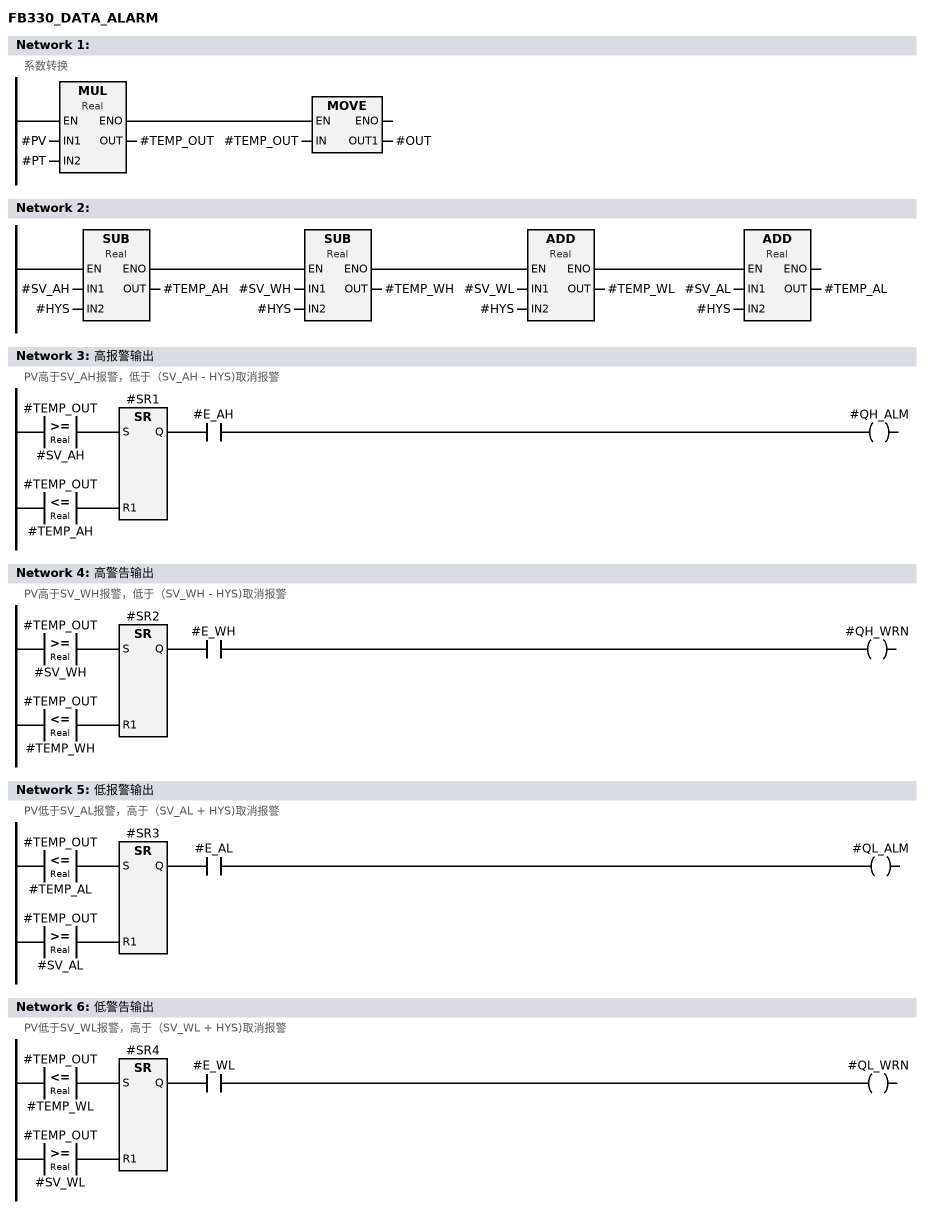
   RUNG wire#powerrail
      { S7_Templates := "SrcType := Real"; S7_GenerateENO := "TRUE" } Mul(in1 := #PV, in2 := #PT, out => #TEMP_OUT)
      { S7_GenerateENO := "TRUE" } Move(in := #TEMP_OUT, out1 => #OUT)
   END_RUNG
   // the same network as SCL:
   // ENO of a box is taken as its EN; it also drops when the box reports an error
   #TEMP_OUT := #PV * #PT;
   #OUT := #TEMP_OUT;
END_REGION

REGION Network 2
   RUNG wire#powerrail
      { S7_Templates := "SrcType := Real"; S7_GenerateENO := "TRUE" } Sub(in1 := #SV_AH, in2 := #HYS, out => #TEMP_AH)
      { S7_Templates := "SrcType := Real"; S7_GenerateENO := "TRUE" } Sub(in1 := #SV_WH, in2 := #HYS, out => #TEMP_WH)
      { S7_Templates := "SrcType := Real"; S7_GenerateENO := "TRUE" } Add(in1 := #SV_WL, in2 := #HYS, out => #TEMP_WL)
      { S7_Templates := "SrcType := Real"; S7_GenerateENO := "TRUE" } Add(in1 := #SV_AL, in2 := #HYS, out => #TEMP_AL)
   END_RUNG
   // the same network as SCL:
   // ENO of a box is taken as its EN; it also drops when the box reports an error
   #TEMP_AH := #SV_AH - #HYS;
   #TEMP_WH := #SV_WH - #HYS;
   #TEMP_WL := #SV_WL + #HYS;
   #TEMP_AL := #SV_AL + #HYS;
END_REGION

REGION Network 3: 高报警输出
   // PV高于SV_AH报警，低于（SV_AH - HYS)取消报警
   RUNG wire#powerrail
      { S7_Templates := "SrcType := Real" } GE_Contact(in1 := #TEMP_OUT, in2 := #SV_AH)
      S_SR(operand := #SR1, r1 := wire#w1)
      Contact( #E_AH )
      Coil( #QH_ALM )
   END_RUNG
   RUNG wire#powerrail
      { S7_Templates := "SrcType := Real" } LE_Contact(in1 := #TEMP_OUT, in2 := #TEMP_AH)
   END_RUNG wire#w1
   // the same network as SCL:
   IF #TEMP_OUT >= #SV_AH THEN
       #SR1 := TRUE;   // SR flip-flop
   END_IF;
   IF #TEMP_OUT <= #TEMP_AH THEN #SR1 := FALSE; END_IF;
   #QH_ALM := #SR1 AND #E_AH;
END_REGION

REGION Network 4: 高警告输出
   // PV高于SV_WH报警，低于（SV_WH - HYS)取消报警
   RUNG wire#powerrail
      { S7_Templates := "SrcType := Real" } GE_Contact(in1 := #TEMP_OUT, in2 := #SV_WH)
      S_SR(operand := #SR2, r1 := wire#w1)
      Contact( #E_WH )
      Coil( #QH_WRN )
   END_RUNG
   RUNG wire#powerrail
      { S7_Templates := "SrcType := Real" } LE_Contact(in1 := #TEMP_OUT, in2 := #TEMP_WH)
   END_RUNG wire#w1
   // the same network as SCL:
   IF #TEMP_OUT >= #SV_WH THEN
       #SR2 := TRUE;   // SR flip-flop
   END_IF;
   IF #TEMP_OUT <= #TEMP_WH THEN #SR2 := FALSE; END_IF;
   #QH_WRN := #SR2 AND #E_WH;
END_REGION

REGION Network 5: 低报警输出
   // PV低于SV_AL报警，高于（SV_AL + HYS)取消报警
   RUNG wire#powerrail
      { S7_Templates := "SrcType := Real" } LE_Contact(in1 := #TEMP_OUT, in2 := #TEMP_AL)
      S_SR(operand := #SR3, r1 := wire#w1)
      Contact( #E_AL )
      Coil( #QL_ALM )
   END_RUNG
   RUNG wire#powerrail
      { S7_Templates := "SrcType := Real" } GE_Contact(in1 := #TEMP_OUT, in2 := #SV_AL)
   END_RUNG wire#w1
   // the same network as SCL:
   IF #TEMP_OUT <= #TEMP_AL THEN
       #SR3 := TRUE;   // SR flip-flop
   END_IF;
   IF #TEMP_OUT >= #SV_AL THEN #SR3 := FALSE; END_IF;
   #QL_ALM := #SR3 AND #E_AL;
END_REGION

REGION Network 6: 低警告输出
   // PV低于SV_WL报警，高于（SV_WL + HYS)取消报警
   RUNG wire#powerrail
      { S7_Templates := "SrcType := Real" } LE_Contact(in1 := #TEMP_OUT, in2 := #TEMP_WL)
      S_SR(operand := #SR4, r1 := wire#w1)
      Contact( #E_WL )
      Coil( #QL_WRN )
   END_RUNG
   RUNG wire#powerrail
      { S7_Templates := "SrcType := Real" } GE_Contact(in1 := #TEMP_OUT, in2 := #SV_WL)
   END_RUNG wire#w1
   // the same network as SCL:
   IF #TEMP_OUT <= #TEMP_WL THEN
       #SR4 := TRUE;   // SR flip-flop
   END_IF;
   IF #TEMP_OUT >= #SV_WL THEN #SR4 := FALSE; END_IF;
   #QL_WRN := #SR4 AND #E_WL;
END_REGION
END_FUNCTION_BLOCK

FUNCTION "电机控制" : Void   // FC1, LAD
{ S7_Optimized_Access := 'FALSE' }
VERSION : 0.1
   VAR_TEMP   // added for the SCL form of the ladder/FBD networks
      _w1 : Bool;
      _s5time1 : S5Time;
      _w2 : Bool;
   END_VAR
BEGIN

REGION Network 1
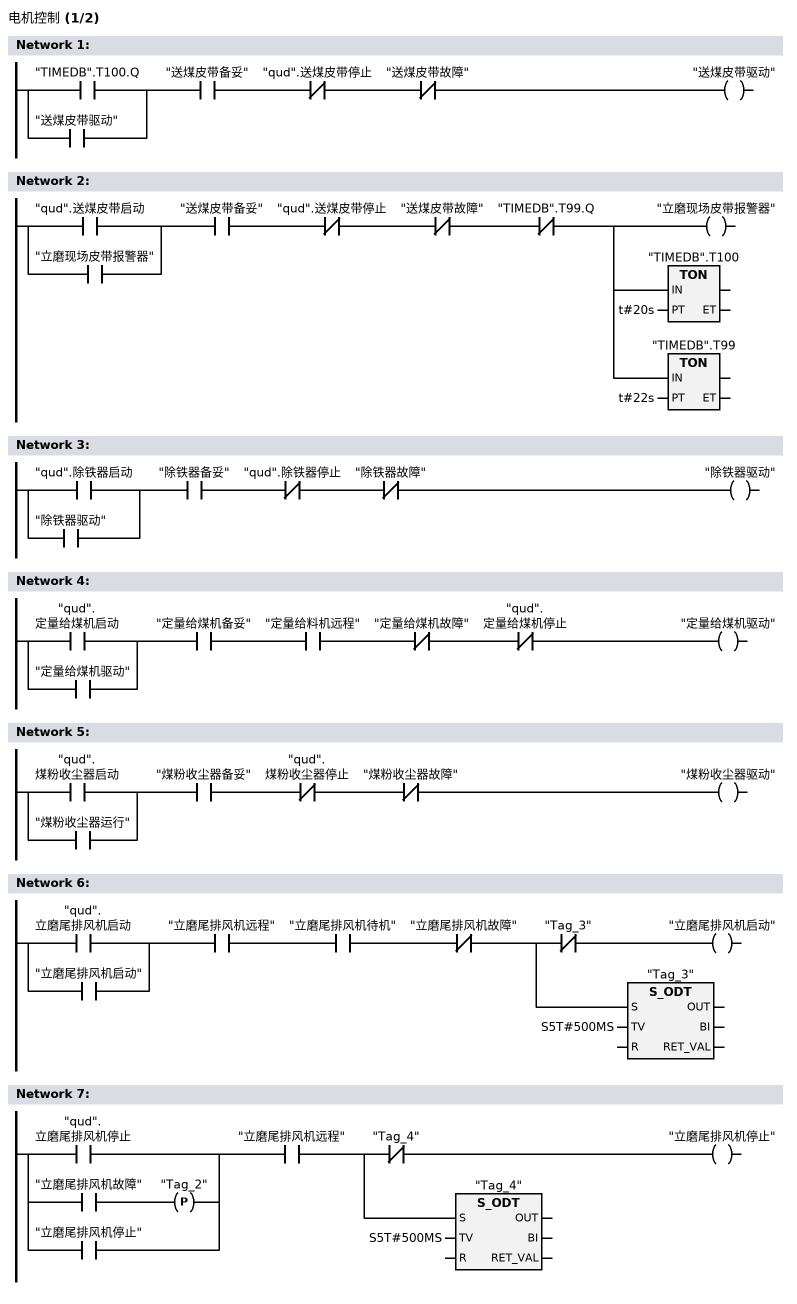
   RUNG wire#powerrail
      Contact( "TIMEDB".T100.Q )
      wire#w1
      Contact( "送煤皮带备妥" )
      I_Contact( "qud".送煤皮带停止 )
      I_Contact( "送煤皮带故障" )
      Coil( "送煤皮带驱动" )
   END_RUNG
   RUNG wire#powerrail
      Contact( "送煤皮带驱动" )
   END_RUNG wire#w1
   // the same network as SCL:
   "送煤皮带驱动" := ("TIMEDB".T100.Q OR "送煤皮带驱动") AND "送煤皮带备妥" AND NOT "qud".送煤皮带停止 AND NOT "送煤皮带故障";
END_REGION

REGION Network 2
   "立磨现场皮带报警器" := ("qud".送煤皮带启动 OR "立磨现场皮带报警器") AND "送煤皮带备妥" AND NOT "qud".送煤皮带停止 AND NOT "送煤皮带故障" AND NOT "TIMEDB".T99.Q;
   "TIMEDB".T100.TON(IN := "立磨现场皮带报警器", PT := t#20s);
   "TIMEDB".T99.TON(IN := "立磨现场皮带报警器", PT := t#22s);
END_REGION

REGION Network 3
   RUNG wire#powerrail
      Contact( "qud".除铁器启动 )
      wire#w1
      Contact( "除铁器备妥" )
      I_Contact( "qud".除铁器停止 )
      I_Contact( "除铁器故障" )
      Coil( "除铁器驱动" )
   END_RUNG
   RUNG wire#powerrail
      Contact( "除铁器驱动" )
   END_RUNG wire#w1
   // the same network as SCL:
   "除铁器驱动" := ("qud".除铁器启动 OR "除铁器驱动") AND "除铁器备妥" AND NOT "qud".除铁器停止 AND NOT "除铁器故障";
END_REGION

REGION Network 4
   RUNG wire#powerrail
      Contact( "qud".定量给煤机启动 )
      wire#w1
      Contact( "定量给煤机备妥" )
      Contact( "定量给料机远程" )
      I_Contact( "定量给煤机故障" )
      I_Contact( "qud".定量给煤机停止 )
      Coil( "定量给煤机驱动" )
   END_RUNG
   RUNG wire#powerrail
      Contact( "定量给煤机驱动" )
   END_RUNG wire#w1
   // the same network as SCL:
   "定量给煤机驱动" := ("qud".定量给煤机启动 OR "定量给煤机驱动") AND "定量给煤机备妥" AND "定量给料机远程" AND NOT "定量给煤机故障" AND NOT "qud".定量给煤机停止;
END_REGION

REGION Network 5
   RUNG wire#powerrail
      Contact( "qud".煤粉收尘器启动 )
      wire#w1
      Contact( "煤粉收尘器备妥" )
      I_Contact( "qud".煤粉收尘器停止 )
      I_Contact( "煤粉收尘器故障" )
      Coil( "煤粉收尘器驱动" )
   END_RUNG
   RUNG wire#powerrail
      Contact( "煤粉收尘器运行" )
   END_RUNG wire#w1
   // the same network as SCL:
   "煤粉收尘器驱动" := ("qud".煤粉收尘器启动 OR "煤粉收尘器运行") AND "煤粉收尘器备妥" AND NOT "qud".煤粉收尘器停止 AND NOT "煤粉收尘器故障";
END_REGION

REGION Network 6
   RUNG wire#powerrail
      Contact( "qud".立磨尾排风机启动 )
      wire#w1
      Contact( "立磨尾排风机远程" )
      Contact( "立磨尾排风机待机" )
      I_Contact( "立磨尾排风机故障" )
      wire#w2
      I_Contact( "Tag_3" )
      Coil( "立磨尾排风机启动" )
   END_RUNG
   RUNG wire#powerrail
      Contact( "立磨尾排风机启动" )
   END_RUNG wire#w1
   RUNG wire#w2
      S_ODT(T_NO := "Tag_3", TV := S5T#500MS, R :=, BI =>, RET_VAL =>)
   END_RUNG
   // the same network as SCL:
   #_w1 := ("qud".立磨尾排风机启动 OR "立磨尾排风机启动") AND "立磨尾排风机远程" AND "立磨尾排风机待机" AND NOT "立磨尾排风机故障";
   "立磨尾排风机启动" := #_w1 AND NOT "Tag_3";
   #_s5time1 := S_ODT(T_NO := "Tag_3", S := #_w1, TV := S5T#500MS);
END_REGION

REGION Network 7
   RUNG wire#powerrail
      Contact( "qud".立磨尾排风机停止 )
      wire#w1
      Contact( "立磨尾排风机远程" )
      wire#w2
      I_Contact( "Tag_4" )
      Coil( "立磨尾排风机停止" )
   END_RUNG
   RUNG wire#powerrail
      Contact( "立磨尾排风机故障" )
      P_Trig( "Tag_2" )
   END_RUNG wire#w1
   RUNG wire#powerrail
      Contact( "立磨尾排风机停止" )
   END_RUNG wire#w1
   RUNG wire#w2
      S_ODT(T_NO := "Tag_4", TV := S5T#500MS, R :=, BI =>, RET_VAL =>)
   END_RUNG
   // the same network as SCL:
   #_w1 := "立磨尾排风机故障" AND NOT "Tag_2";   // rising edge
   "Tag_2" := "立磨尾排风机故障";
   #_w2 := ("qud".立磨尾排风机停止 OR #_w1 OR "立磨尾排风机停止") AND "立磨尾排风机远程";
   "立磨尾排风机停止" := #_w2 AND NOT "Tag_4";
   #_s5time1 := S_ODT(T_NO := "Tag_4", S := #_w2, TV := S5T#500MS);
END_REGION

REGION Network 8
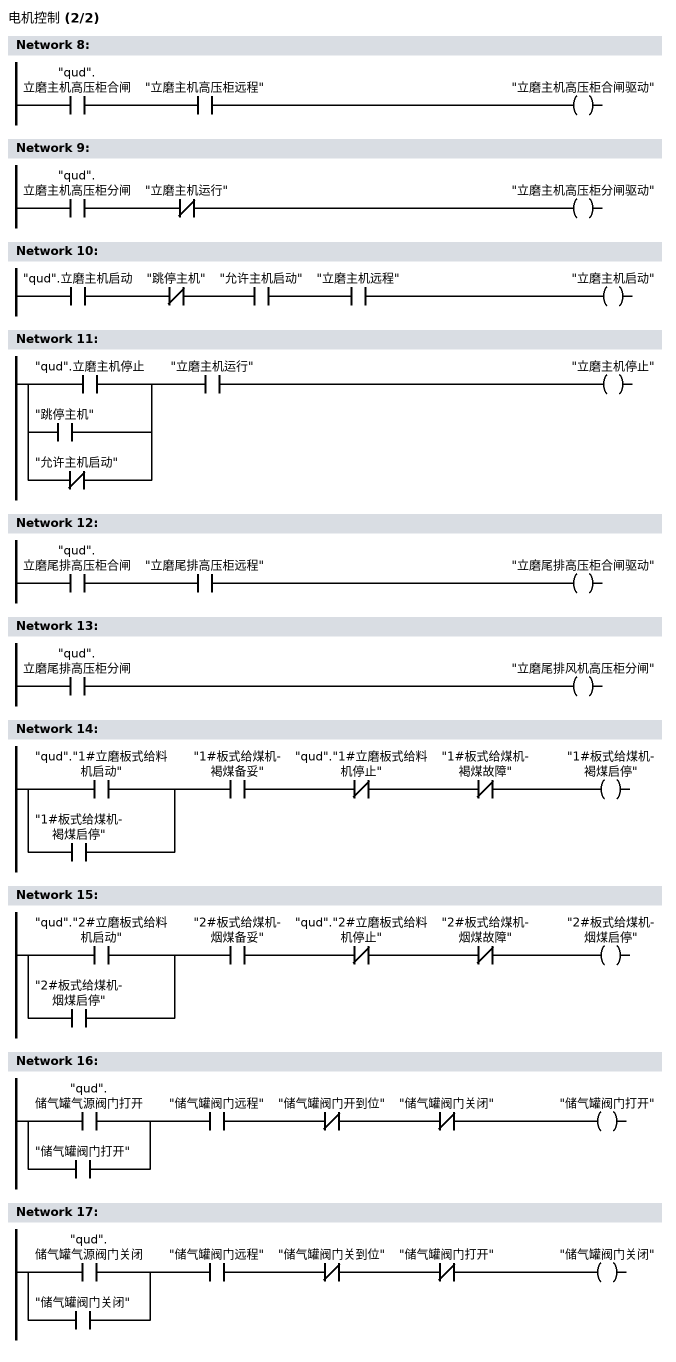
   RUNG wire#powerrail
      Contact( "qud".立磨主机高压柜合闸 )
      Contact( "立磨主机高压柜远程" )
      Coil( "立磨主机高压柜合闸驱动" )
   END_RUNG
   // the same network as SCL:
   "立磨主机高压柜合闸驱动" := "qud".立磨主机高压柜合闸 AND "立磨主机高压柜远程";
END_REGION

REGION Network 9
   RUNG wire#powerrail
      Contact( "qud".立磨主机高压柜分闸 )
      I_Contact( "立磨主机运行" )
      Coil( "立磨主机高压柜分闸驱动" )
   END_RUNG
   // the same network as SCL:
   "立磨主机高压柜分闸驱动" := "qud".立磨主机高压柜分闸 AND NOT "立磨主机运行";
END_REGION

REGION Network 10
   RUNG wire#powerrail
      Contact( "qud".立磨主机启动 )
      I_Contact( "跳停主机" )
      Contact( "允许主机启动" )
      Contact( "立磨主机远程" )
      Coil( "立磨主机启动" )
   END_RUNG
   // the same network as SCL:
   "立磨主机启动" := "qud".立磨主机启动 AND NOT "跳停主机" AND "允许主机启动" AND "立磨主机远程";
END_REGION

REGION Network 11
   RUNG wire#powerrail
      Contact( "qud".立磨主机停止 )
      wire#w1
      Contact( "立磨主机运行" )
      Coil( "立磨主机停止" )
   END_RUNG
   RUNG wire#powerrail
      Contact( "跳停主机" )
   END_RUNG wire#w1
   RUNG wire#powerrail
      I_Contact( "允许主机启动" )
   END_RUNG wire#w1
   // the same network as SCL:
   "立磨主机停止" := ("qud".立磨主机停止 OR "跳停主机" OR NOT "允许主机启动") AND "立磨主机运行";
END_REGION

REGION Network 12
   RUNG wire#powerrail
      Contact( "qud".立磨尾排高压柜合闸 )
      Contact( "立磨尾排高压柜远程" )
      Coil( "立磨尾排高压柜合闸驱动" )
   END_RUNG
   // the same network as SCL:
   "立磨尾排高压柜合闸驱动" := "qud".立磨尾排高压柜合闸 AND "立磨尾排高压柜远程";
END_REGION

REGION Network 13
   RUNG wire#powerrail
      Contact( "qud".立磨尾排高压柜分闸 )
      Coil( "立磨尾排风机高压柜分闸" )
   END_RUNG
   // the same network as SCL:
   "立磨尾排风机高压柜分闸" := "qud".立磨尾排高压柜分闸;
END_REGION

REGION Network 14
   RUNG wire#powerrail
      Contact( "qud"."1#立磨板式给料机启动" )
      wire#w1
      Contact( "1#板式给煤机-褐煤备妥" )
      I_Contact( "qud"."1#立磨板式给料机停止" )
      I_Contact( "1#板式给煤机-褐煤故障" )
      Coil( "1#板式给煤机-褐煤启停" )
   END_RUNG
   RUNG wire#powerrail
      Contact( "1#板式给煤机-褐煤启停" )
   END_RUNG wire#w1
   // the same network as SCL:
   "1#板式给煤机-褐煤启停" := ("qud"."1#立磨板式给料机启动" OR "1#板式给煤机-褐煤启停") AND "1#板式给煤机-褐煤备妥" AND NOT "qud"."1#立磨板式给料机停止" AND NOT "1#板式给煤机-褐煤故障";
END_REGION

REGION Network 15
   RUNG wire#powerrail
      Contact( "qud"."2#立磨板式给料机启动" )
      wire#w1
      Contact( "2#板式给煤机-烟煤备妥" )
      I_Contact( "qud"."2#立磨板式给料机停止" )
      I_Contact( "2#板式给煤机-烟煤故障" )
      Coil( "2#板式给煤机-烟煤启停" )
   END_RUNG
   RUNG wire#powerrail
      Contact( "2#板式给煤机-烟煤启停" )
   END_RUNG wire#w1
   // the same network as SCL:
   "2#板式给煤机-烟煤启停" := ("qud"."2#立磨板式给料机启动" OR "2#板式给煤机-烟煤启停") AND "2#板式给煤机-烟煤备妥" AND NOT "qud"."2#立磨板式给料机停止" AND NOT "2#板式给煤机-烟煤故障";
END_REGION

REGION Network 16
   RUNG wire#powerrail
      Contact( "qud".储气罐气源阀门打开 )
      wire#w1
      Contact( "储气罐阀门远程" )
      I_Contact( "储气罐阀门开到位" )
      I_Contact( "储气罐阀门关闭" )
      Coil( "储气罐阀门打开" )
   END_RUNG
   RUNG wire#powerrail
      Contact( "储气罐阀门打开" )
   END_RUNG wire#w1
   // the same network as SCL:
   "储气罐阀门打开" := ("qud".储气罐气源阀门打开 OR "储气罐阀门打开") AND "储气罐阀门远程" AND NOT "储气罐阀门开到位" AND NOT "储气罐阀门关闭";
END_REGION

REGION Network 17
   RUNG wire#powerrail
      Contact( "qud".储气罐气源阀门关闭 )
      wire#w1
      Contact( "储气罐阀门远程" )
      I_Contact( "储气罐阀门关到位" )
      I_Contact( "储气罐阀门打开" )
      Coil( "储气罐阀门关闭" )
   END_RUNG
   RUNG wire#powerrail
      Contact( "储气罐阀门关闭" )
   END_RUNG wire#w1
   // the same network as SCL:
   "储气罐阀门关闭" := ("qud".储气罐气源阀门关闭 OR "储气罐阀门关闭") AND "储气罐阀门远程" AND NOT "储气罐阀门关到位" AND NOT "储气罐阀门打开";
END_REGION
END_FUNCTION

FUNCTION "模拟量" : Void   // FC2, LAD
{ S7_Optimized_Access := 'FALSE' }
VERSION : 0.1
BEGIN

REGION Network 1
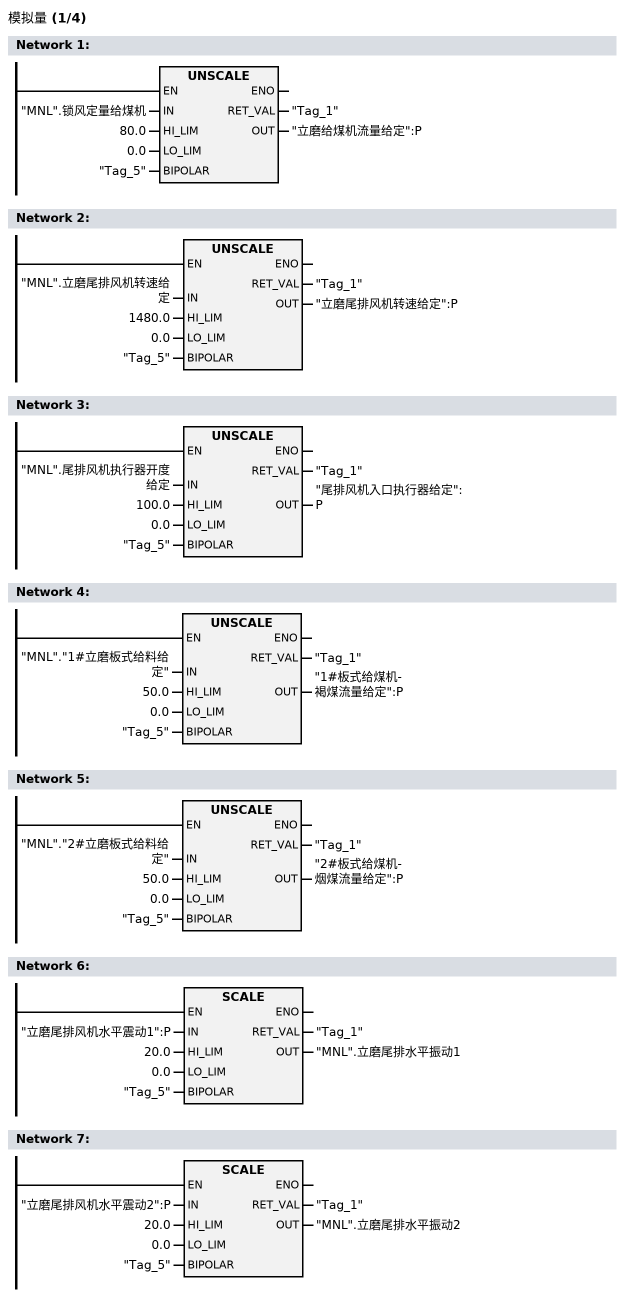
   "Tag_1" := UNSCALE(IN := "MNL".锁风定量给煤机,
                      HI_LIM := 80.0,
                      LO_LIM := 0.0,
                      BIPOLAR := "Tag_5",
                      OUT => "立磨给煤机流量给定":P);
END_REGION

REGION Network 2
   "Tag_1" := UNSCALE(IN := "MNL".立磨尾排风机转速给定,
                      HI_LIM := 1480.0,
                      LO_LIM := 0.0,
                      BIPOLAR := "Tag_5",
                      OUT => "立磨尾排风机转速给定":P);
END_REGION

REGION Network 3
   "Tag_1" := UNSCALE(IN := "MNL".尾排风机执行器开度给定,
                      HI_LIM := 100.0,
                      LO_LIM := 0.0,
                      BIPOLAR := "Tag_5",
                      OUT => "尾排风机入口执行器给定":P);
END_REGION

REGION Network 4
   "Tag_1" := UNSCALE(IN := "MNL"."1#立磨板式给料给定",
                      HI_LIM := 50.0,
                      LO_LIM := 0.0,
                      BIPOLAR := "Tag_5",
                      OUT => "1#板式给煤机-褐煤流量给定":P);
END_REGION

REGION Network 5
   "Tag_1" := UNSCALE(IN := "MNL"."2#立磨板式给料给定",
                      HI_LIM := 50.0,
                      LO_LIM := 0.0,
                      BIPOLAR := "Tag_5",
                      OUT => "2#板式给煤机-烟煤流量给定":P);
END_REGION

REGION Network 6
   "Tag_1" := SCALE(IN := "立磨尾排风机水平震动1":P,
                    HI_LIM := 20.0,
                    LO_LIM := 0.0,
                    BIPOLAR := "Tag_5",
                    OUT => "MNL".立磨尾排水平振动1);
END_REGION

REGION Network 7
   "Tag_1" := SCALE(IN := "立磨尾排风机水平震动2":P,
                    HI_LIM := 20.0,
                    LO_LIM := 0.0,
                    BIPOLAR := "Tag_5",
                    OUT => "MNL".立磨尾排水平振动2);
END_REGION

REGION Network 8
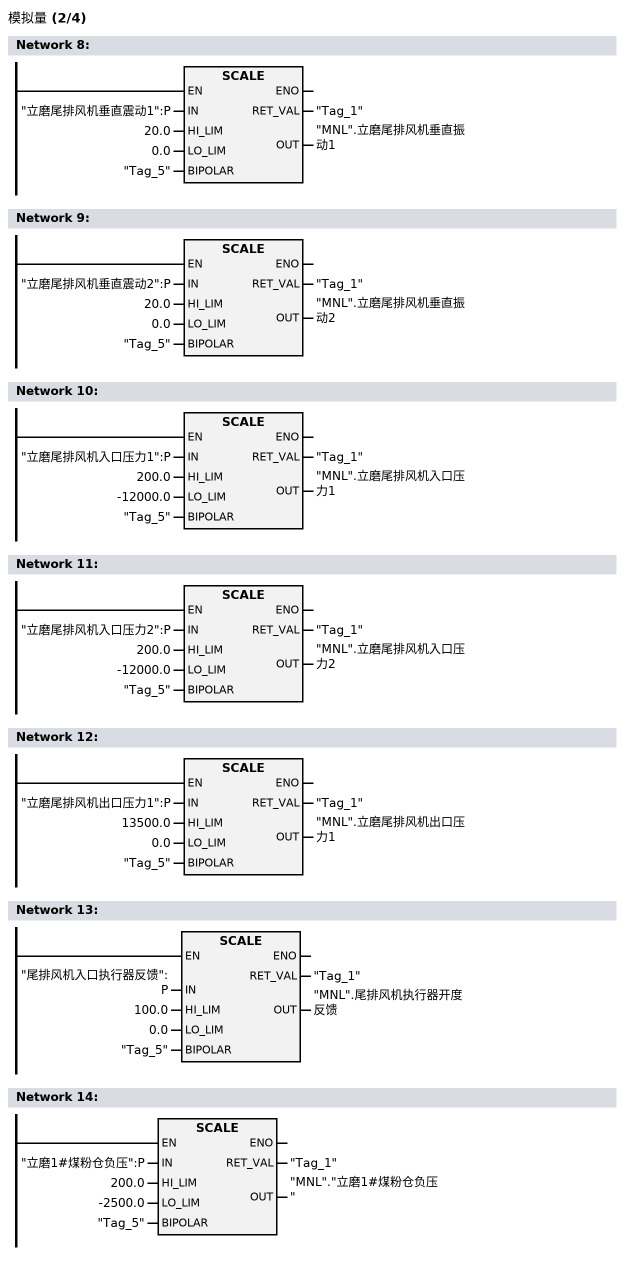
   "Tag_1" := SCALE(IN := "立磨尾排风机垂直震动1":P,
                    HI_LIM := 20.0,
                    LO_LIM := 0.0,
                    BIPOLAR := "Tag_5",
                    OUT => "MNL".立磨尾排风机垂直振动1);
END_REGION

REGION Network 9
   "Tag_1" := SCALE(IN := "立磨尾排风机垂直震动2":P,
                    HI_LIM := 20.0,
                    LO_LIM := 0.0,
                    BIPOLAR := "Tag_5",
                    OUT => "MNL".立磨尾排风机垂直振动2);
END_REGION

REGION Network 10
   "Tag_1" := SCALE(IN := "立磨尾排风机入口压力1":P,
                    HI_LIM := 200.0,
                    LO_LIM := -12000.0,
                    BIPOLAR := "Tag_5",
                    OUT => "MNL".立磨尾排风机入口压力1);
END_REGION

REGION Network 11
   "Tag_1" := SCALE(IN := "立磨尾排风机入口压力2":P,
                    HI_LIM := 200.0,
                    LO_LIM := -12000.0,
                    BIPOLAR := "Tag_5",
                    OUT => "MNL".立磨尾排风机入口压力2);
END_REGION

REGION Network 12
   "Tag_1" := SCALE(IN := "立磨尾排风机出口压力1":P,
                    HI_LIM := 13500.0,
                    LO_LIM := 0.0,
                    BIPOLAR := "Tag_5",
                    OUT => "MNL".立磨尾排风机出口压力1);
END_REGION

REGION Network 13
   "Tag_1" := SCALE(IN := "尾排风机入口执行器反馈":P,
                    HI_LIM := 100.0,
                    LO_LIM := 0.0,
                    BIPOLAR := "Tag_5",
                    OUT => "MNL".尾排风机执行器开度反馈);
END_REGION

REGION Network 14
   "Tag_1" := SCALE(IN := "立磨1#煤粉仓负压":P,
                    HI_LIM := 200.0,
                    LO_LIM := -2500.0,
                    BIPOLAR := "Tag_5",
                    OUT => "MNL"."立磨1#煤粉仓负压");
END_REGION

REGION Network 15
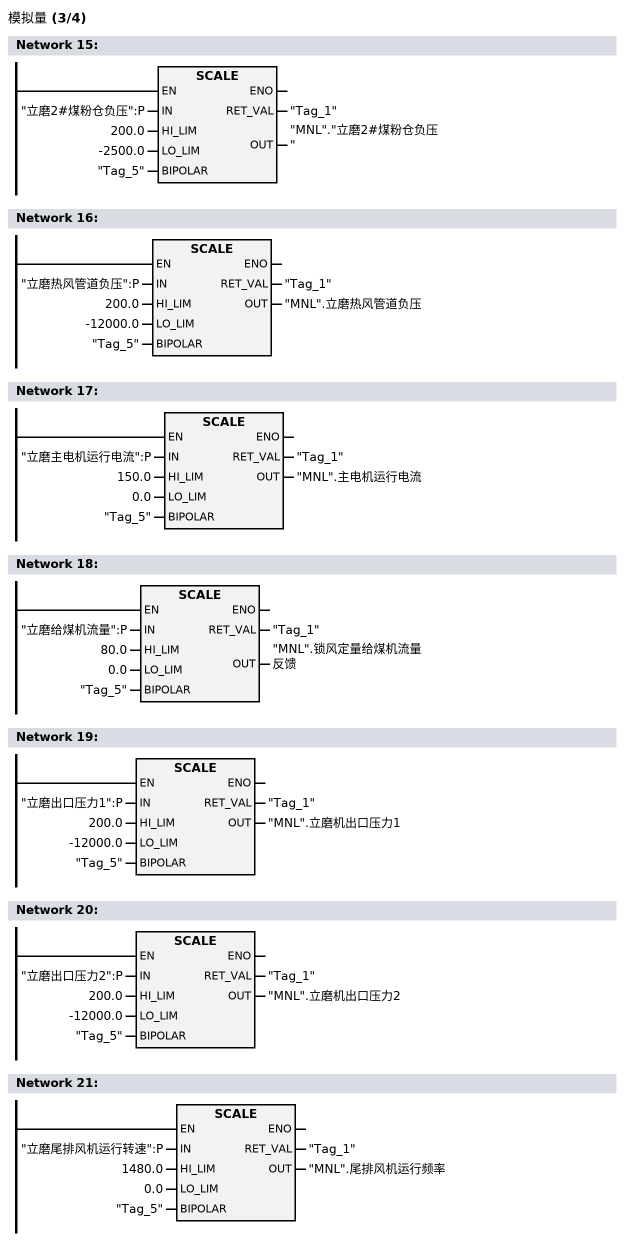
   "Tag_1" := SCALE(IN := "立磨2#煤粉仓负压":P,
                    HI_LIM := 200.0,
                    LO_LIM := -2500.0,
                    BIPOLAR := "Tag_5",
                    OUT => "MNL"."立磨2#煤粉仓负压");
END_REGION

REGION Network 16
   "Tag_1" := SCALE(IN := "立磨热风管道负压":P,
                    HI_LIM := 200.0,
                    LO_LIM := -12000.0,
                    BIPOLAR := "Tag_5",
                    OUT => "MNL".立磨热风管道负压);
END_REGION

REGION Network 17
   "Tag_1" := SCALE(IN := "立磨主电机运行电流":P,
                    HI_LIM := 150.0,
                    LO_LIM := 0.0,
                    BIPOLAR := "Tag_5",
                    OUT => "MNL".主电机运行电流);
END_REGION

REGION Network 18
   "Tag_1" := SCALE(IN := "立磨给煤机流量":P,
                    HI_LIM := 80.0,
                    LO_LIM := 0.0,
                    BIPOLAR := "Tag_5",
                    OUT => "MNL".锁风定量给煤机流量反馈);
END_REGION

REGION Network 19
   "Tag_1" := SCALE(IN := "立磨出口压力1":P,
                    HI_LIM := 200.0,
                    LO_LIM := -12000.0,
                    BIPOLAR := "Tag_5",
                    OUT => "MNL".立磨机出口压力1);
END_REGION

REGION Network 20
   "Tag_1" := SCALE(IN := "立磨出口压力2":P,
                    HI_LIM := 200.0,
                    LO_LIM := -12000.0,
                    BIPOLAR := "Tag_5",
                    OUT => "MNL".立磨机出口压力2);
END_REGION

REGION Network 21
   "Tag_1" := SCALE(IN := "立磨尾排风机运行转速":P,
                    HI_LIM := 1480.0,
                    LO_LIM := 0.0,
                    BIPOLAR := "Tag_5",
                    OUT => "MNL".尾排风机运行频率);
END_REGION

REGION Network 22
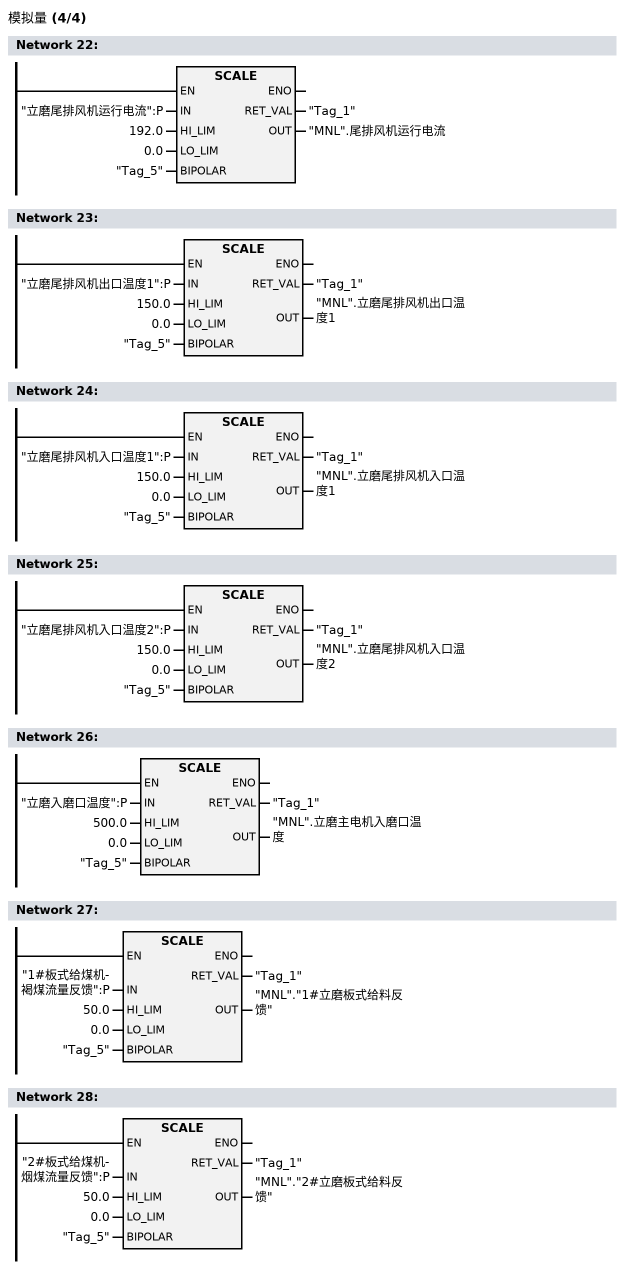
   "Tag_1" := SCALE(IN := "立磨尾排风机运行电流":P,
                    HI_LIM := 192.0,
                    LO_LIM := 0.0,
                    BIPOLAR := "Tag_5",
                    OUT => "MNL".尾排风机运行电流);
END_REGION

REGION Network 23
   "Tag_1" := SCALE(IN := "立磨尾排风机出口温度1":P,
                    HI_LIM := 150.0,
                    LO_LIM := 0.0,
                    BIPOLAR := "Tag_5",
                    OUT => "MNL".立磨尾排风机出口温度1);
END_REGION

REGION Network 24
   "Tag_1" := SCALE(IN := "立磨尾排风机入口温度1":P,
                    HI_LIM := 150.0,
                    LO_LIM := 0.0,
                    BIPOLAR := "Tag_5",
                    OUT => "MNL".立磨尾排风机入口温度1);
END_REGION

REGION Network 25
   "Tag_1" := SCALE(IN := "立磨尾排风机入口温度2":P,
                    HI_LIM := 150.0,
                    LO_LIM := 0.0,
                    BIPOLAR := "Tag_5",
                    OUT => "MNL".立磨尾排风机入口温度2);
END_REGION

REGION Network 26
   "Tag_1" := SCALE(IN := "立磨入磨口温度":P,
                    HI_LIM := 500.0,
                    LO_LIM := 0.0,
                    BIPOLAR := "Tag_5",
                    OUT => "MNL".立磨主电机入磨口温度);
END_REGION

REGION Network 27
   "Tag_1" := SCALE(IN := "1#板式给煤机-褐煤流量反馈":P,
                    HI_LIM := 50.0,
                    LO_LIM := 0.0,
                    BIPOLAR := "Tag_5",
                    OUT => "MNL"."1#立磨板式给料反馈");
END_REGION

REGION Network 28
   "Tag_1" := SCALE(IN := "2#板式给煤机-烟煤流量反馈":P,
                    HI_LIM := 50.0,
                    LO_LIM := 0.0,
                    BIPOLAR := "Tag_5",
                    OUT => "MNL"."2#立磨板式给料反馈");
END_REGION
END_FUNCTION

FUNCTION "仪表数据" : Void   // FC4, LAD
{ S7_Optimized_Access := 'FALSE' }
VERSION : 0.1
BEGIN

REGION Network 1
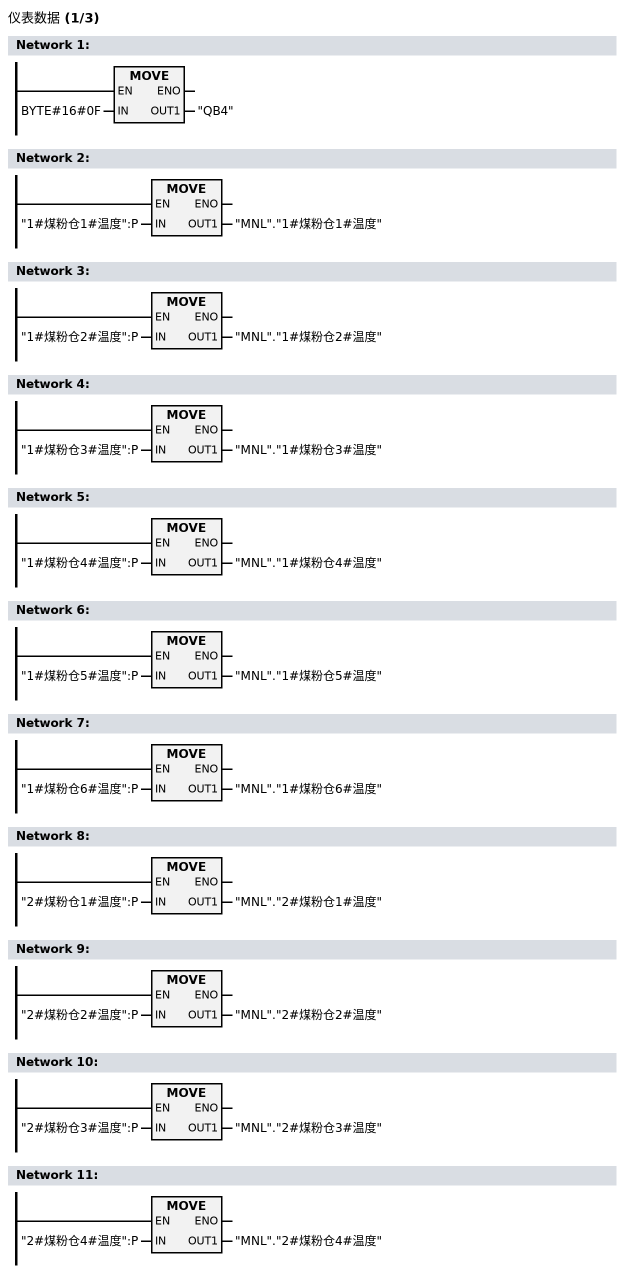
   RUNG wire#powerrail
      { S7_GenerateENO := "TRUE" } Move(in := BYTE#16#0F, out1 => "QB4")
   END_RUNG
   // the same network as SCL:
   "QB4" := BYTE#16#0F;
END_REGION

REGION Network 2
   RUNG wire#powerrail
      { S7_GenerateENO := "TRUE" } Move(in := "1#煤粉仓1#温度":P, out1 => "MNL"."1#煤粉仓1#温度")
   END_RUNG
   // the same network as SCL:
   "MNL"."1#煤粉仓1#温度" := "1#煤粉仓1#温度":P;
END_REGION

REGION Network 3
   RUNG wire#powerrail
      { S7_GenerateENO := "TRUE" } Move(in := "1#煤粉仓2#温度":P, out1 => "MNL"."1#煤粉仓2#温度")
   END_RUNG
   // the same network as SCL:
   "MNL"."1#煤粉仓2#温度" := "1#煤粉仓2#温度":P;
END_REGION

REGION Network 4
   RUNG wire#powerrail
      { S7_GenerateENO := "TRUE" } Move(in := "1#煤粉仓3#温度":P, out1 => "MNL"."1#煤粉仓3#温度")
   END_RUNG
   // the same network as SCL:
   "MNL"."1#煤粉仓3#温度" := "1#煤粉仓3#温度":P;
END_REGION

REGION Network 5
   RUNG wire#powerrail
      { S7_GenerateENO := "TRUE" } Move(in := "1#煤粉仓4#温度":P, out1 => "MNL"."1#煤粉仓4#温度")
   END_RUNG
   // the same network as SCL:
   "MNL"."1#煤粉仓4#温度" := "1#煤粉仓4#温度":P;
END_REGION

REGION Network 6
   RUNG wire#powerrail
      { S7_GenerateENO := "TRUE" } Move(in := "1#煤粉仓5#温度":P, out1 => "MNL"."1#煤粉仓5#温度")
   END_RUNG
   // the same network as SCL:
   "MNL"."1#煤粉仓5#温度" := "1#煤粉仓5#温度":P;
END_REGION

REGION Network 7
   RUNG wire#powerrail
      { S7_GenerateENO := "TRUE" } Move(in := "1#煤粉仓6#温度":P, out1 => "MNL"."1#煤粉仓6#温度")
   END_RUNG
   // the same network as SCL:
   "MNL"."1#煤粉仓6#温度" := "1#煤粉仓6#温度":P;
END_REGION

REGION Network 8
   RUNG wire#powerrail
      { S7_GenerateENO := "TRUE" } Move(in := "2#煤粉仓1#温度":P, out1 => "MNL"."2#煤粉仓1#温度")
   END_RUNG
   // the same network as SCL:
   "MNL"."2#煤粉仓1#温度" := "2#煤粉仓1#温度":P;
END_REGION

REGION Network 9
   RUNG wire#powerrail
      { S7_GenerateENO := "TRUE" } Move(in := "2#煤粉仓2#温度":P, out1 => "MNL"."2#煤粉仓2#温度")
   END_RUNG
   // the same network as SCL:
   "MNL"."2#煤粉仓2#温度" := "2#煤粉仓2#温度":P;
END_REGION

REGION Network 10
   RUNG wire#powerrail
      { S7_GenerateENO := "TRUE" } Move(in := "2#煤粉仓3#温度":P, out1 => "MNL"."2#煤粉仓3#温度")
   END_RUNG
   // the same network as SCL:
   "MNL"."2#煤粉仓3#温度" := "2#煤粉仓3#温度":P;
END_REGION

REGION Network 11
   RUNG wire#powerrail
      { S7_GenerateENO := "TRUE" } Move(in := "2#煤粉仓4#温度":P, out1 => "MNL"."2#煤粉仓4#温度")
   END_RUNG
   // the same network as SCL:
   "MNL"."2#煤粉仓4#温度" := "2#煤粉仓4#温度":P;
END_REGION

REGION Network 12
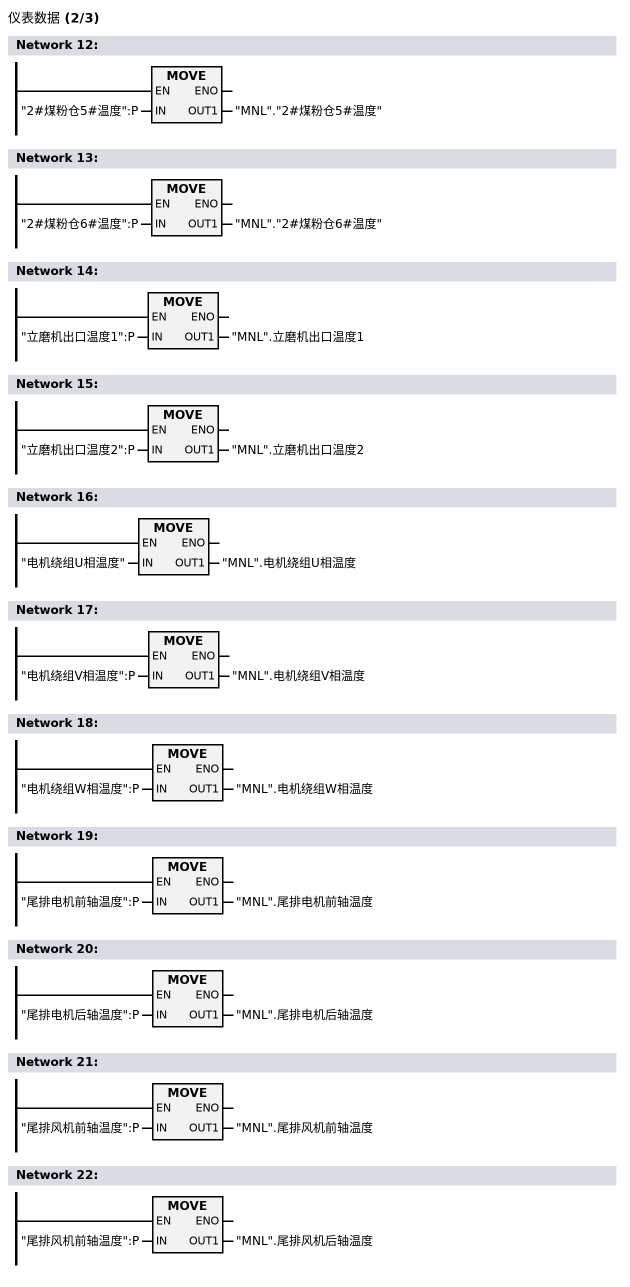
   RUNG wire#powerrail
      { S7_GenerateENO := "TRUE" } Move(in := "2#煤粉仓5#温度":P, out1 => "MNL"."2#煤粉仓5#温度")
   END_RUNG
   // the same network as SCL:
   "MNL"."2#煤粉仓5#温度" := "2#煤粉仓5#温度":P;
END_REGION

REGION Network 13
   RUNG wire#powerrail
      { S7_GenerateENO := "TRUE" } Move(in := "2#煤粉仓6#温度":P, out1 => "MNL"."2#煤粉仓6#温度")
   END_RUNG
   // the same network as SCL:
   "MNL"."2#煤粉仓6#温度" := "2#煤粉仓6#温度":P;
END_REGION

REGION Network 14
   RUNG wire#powerrail
      { S7_GenerateENO := "TRUE" } Move(in := "立磨机出口温度1":P, out1 => "MNL".立磨机出口温度1)
   END_RUNG
   // the same network as SCL:
   "MNL".立磨机出口温度1 := "立磨机出口温度1":P;
END_REGION

REGION Network 15
   RUNG wire#powerrail
      { S7_GenerateENO := "TRUE" } Move(in := "立磨机出口温度2":P, out1 => "MNL".立磨机出口温度2)
   END_RUNG
   // the same network as SCL:
   "MNL".立磨机出口温度2 := "立磨机出口温度2":P;
END_REGION

REGION Network 16
   RUNG wire#powerrail
      { S7_GenerateENO := "TRUE" } Move(in := "电机绕组U相温度", out1 => "MNL".电机绕组U相温度)
   END_RUNG
   // the same network as SCL:
   "MNL".电机绕组U相温度 := "电机绕组U相温度";
END_REGION

REGION Network 17
   RUNG wire#powerrail
      { S7_GenerateENO := "TRUE" } Move(in := "电机绕组V相温度":P, out1 => "MNL".电机绕组V相温度)
   END_RUNG
   // the same network as SCL:
   "MNL".电机绕组V相温度 := "电机绕组V相温度":P;
END_REGION

REGION Network 18
   RUNG wire#powerrail
      { S7_GenerateENO := "TRUE" } Move(in := "电机绕组W相温度":P, out1 => "MNL".电机绕组W相温度)
   END_RUNG
   // the same network as SCL:
   "MNL".电机绕组W相温度 := "电机绕组W相温度":P;
END_REGION

REGION Network 19
   RUNG wire#powerrail
      { S7_GenerateENO := "TRUE" } Move(in := "尾排电机前轴温度":P, out1 => "MNL".尾排电机前轴温度)
   END_RUNG
   // the same network as SCL:
   "MNL".尾排电机前轴温度 := "尾排电机前轴温度":P;
END_REGION

REGION Network 20
   RUNG wire#powerrail
      { S7_GenerateENO := "TRUE" } Move(in := "尾排电机后轴温度":P, out1 => "MNL".尾排电机后轴温度)
   END_RUNG
   // the same network as SCL:
   "MNL".尾排电机后轴温度 := "尾排电机后轴温度":P;
END_REGION

REGION Network 21
   RUNG wire#powerrail
      { S7_GenerateENO := "TRUE" } Move(in := "尾排风机前轴温度":P, out1 => "MNL".尾排风机前轴温度)
   END_RUNG
   // the same network as SCL:
   "MNL".尾排风机前轴温度 := "尾排风机前轴温度":P;
END_REGION

REGION Network 22
   RUNG wire#powerrail
      { S7_GenerateENO := "TRUE" } Move(in := "尾排风机前轴温度":P, out1 => "MNL".尾排风机后轴温度)
   END_RUNG
   // the same network as SCL:
   "MNL".尾排风机后轴温度 := "尾排风机前轴温度":P;
END_REGION

REGION Network 23
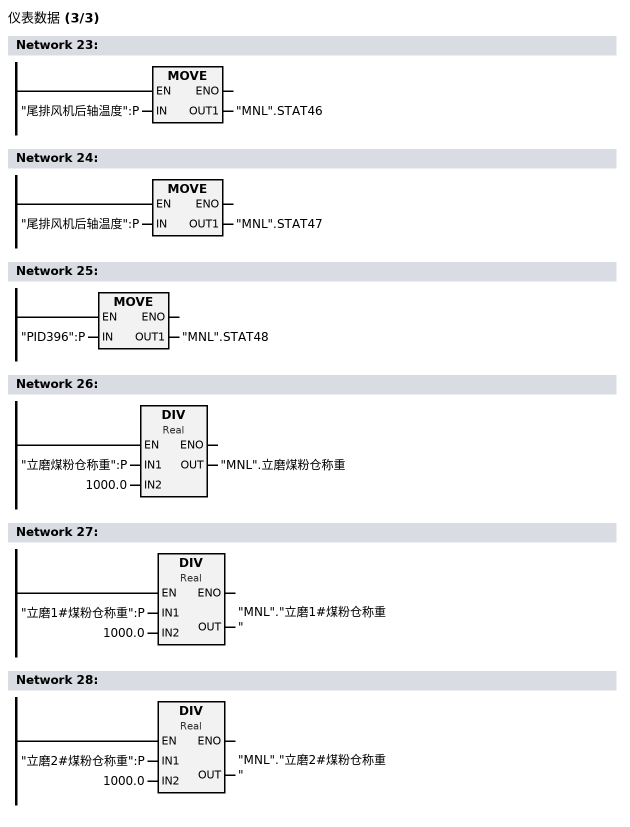
   RUNG wire#powerrail
      { S7_GenerateENO := "TRUE" } Move(in := "尾排风机后轴温度":P, out1 => "MNL".STAT46)
   END_RUNG
   // the same network as SCL:
   "MNL".STAT46 := "尾排风机后轴温度":P;
END_REGION

REGION Network 24
   RUNG wire#powerrail
      { S7_GenerateENO := "TRUE" } Move(in := "尾排风机后轴温度":P, out1 => "MNL".STAT47)
   END_RUNG
   // the same network as SCL:
   "MNL".STAT47 := "尾排风机后轴温度":P;
END_REGION

REGION Network 25
   RUNG wire#powerrail
      { S7_GenerateENO := "TRUE" } Move(in := "PID396":P, out1 => "MNL".STAT48)
   END_RUNG
   // the same network as SCL:
   "MNL".STAT48 := "PID396":P;
END_REGION

REGION Network 26
   RUNG wire#powerrail
      { S7_Templates := "SrcType := Real" } Div(in1 := "立磨煤粉仓称重":P, in2 := 1000.0, out => "MNL".立磨煤粉仓称重)
   END_RUNG
   // the same network as SCL:
   "MNL".立磨煤粉仓称重 := "立磨煤粉仓称重":P / 1000.0;
END_REGION

REGION Network 27
   RUNG wire#powerrail
      { S7_Templates := "SrcType := Real" } Div(in1 := "立磨1#煤粉仓称重":P, in2 := 1000.0, out => "MNL"."立磨1#煤粉仓称重")
   END_RUNG
   // the same network as SCL:
   "MNL"."立磨1#煤粉仓称重" := "立磨1#煤粉仓称重":P / 1000.0;
END_REGION

REGION Network 28
   RUNG wire#powerrail
      { S7_Templates := "SrcType := Real" } Div(in1 := "立磨2#煤粉仓称重":P, in2 := 1000.0, out => "MNL"."立磨2#煤粉仓称重")
   END_RUNG
   // the same network as SCL:
   "MNL"."立磨2#煤粉仓称重" := "立磨2#煤粉仓称重":P / 1000.0;
END_REGION
END_FUNCTION

FUNCTION "温度报警输出" : Void   // FC7, LAD
{ S7_Optimized_Access := 'TRUE' }
VERSION : 0.1
   VAR_TEMP   // added for the SCL form of the ladder/FBD networks
      _w1 : Bool;
   END_VAR
BEGIN

REGION Network 1
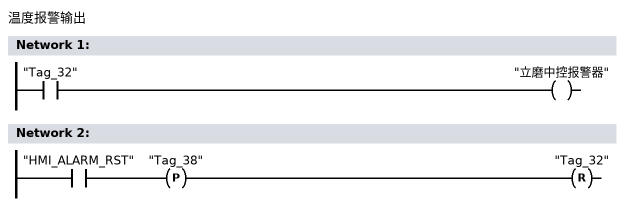
   RUNG wire#powerrail
      Contact( "Tag_32" )
      Coil( "立磨中控报警器" )
   END_RUNG
   // the same network as SCL:
   "立磨中控报警器" := "Tag_32";
END_REGION

REGION Network 2
   RUNG wire#powerrail
      Contact( "HMI_ALARM_RST" )
      P_Trig( "Tag_38" )
      R_Coil( "Tag_32" )
   END_RUNG
   // the same network as SCL:
   #_w1 := "HMI_ALARM_RST" AND NOT "Tag_38";   // rising edge
   "Tag_38" := "HMI_ALARM_RST";
   IF #_w1 THEN "Tag_32" := FALSE; END_IF;
END_REGION
END_FUNCTION

FUNCTION "FC11_DATA_ALARM_FC" : Void   // FC11, LAD
{ S7_Optimized_Access := 'TRUE' }
VERSION : 0.1
   VAR_TEMP   // added for the SCL form of the ladder/FBD networks
      _w1 : Bool;
      _w2 : Bool;
   END_VAR
BEGIN

REGION Network 1
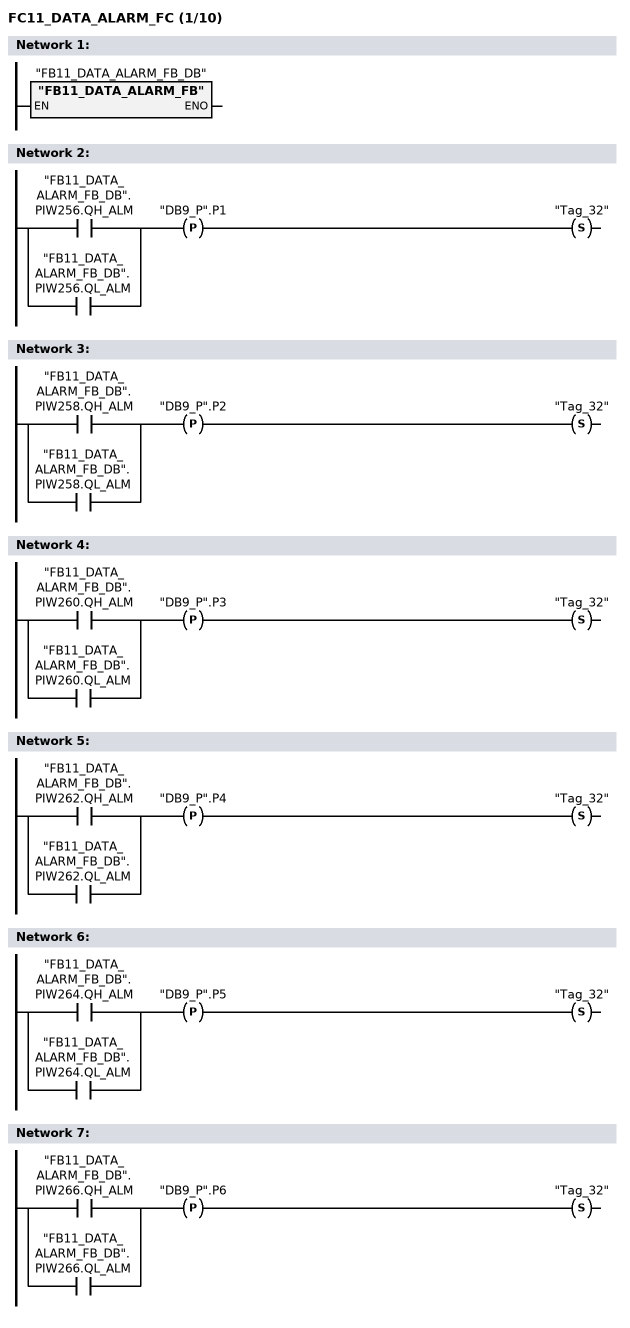
   RUNG wire#powerrail
      "FB11_DATA_ALARM_FB_DB"()
   END_RUNG
   // the same network as SCL:
   "FB11_DATA_ALARM_FB_DB"();   // "FB11_DATA_ALARM_FB"
END_REGION

REGION Network 2
   RUNG wire#powerrail
      Contact( "FB11_DATA_ALARM_FB_DB".PIW256.QH_ALM )
      wire#w1
      P_Trig( "DB9_P".P1 )
      S_Coil( "Tag_32" )
   END_RUNG
   RUNG wire#powerrail
      Contact( "FB11_DATA_ALARM_FB_DB".PIW256.QL_ALM )
   END_RUNG wire#w1
   // the same network as SCL:
   #_w1 := "FB11_DATA_ALARM_FB_DB".PIW256.QH_ALM OR "FB11_DATA_ALARM_FB_DB".PIW256.QL_ALM;
   #_w2 := #_w1 AND NOT "DB9_P".P1;   // rising edge
   "DB9_P".P1 := #_w1;
   IF #_w2 THEN "Tag_32" := TRUE; END_IF;
END_REGION
